// TIA Portal project "HydroPlantProject_V15.1" (V15.1)

(* hardware
DEVICE "S71500/ET200MP station_1"  S7-1500 station
   slot 0: "Rail_0"  Rack  6ES7 590-1***0-0AA0
   slot 1: "PLC_1"  CPU 1511-1 PN  6ES7 511-1AK00-0AB0  V1.8
      slot 3: "CPU display_1"  6ES7591-1AA00-0AA0
DEVICE "PC-System_1"  SIMATIC PC station
   slot 0: "SIMATIC PC station"  Rail  SIMATIC PC-Station  V1.0
      slot 125: "Stationmanager"  Station_Manager  V6.0.4
   slot 1: "HMI_RT_1"  WinCC RT Professional  6AV2 105-0xxxx-xxxx  15.1.0.0
   slot 2: "IE general_1"  IE General  IE_CP  V8.2.0
*)

// ===== PLC "PLC_1"  CPU 1511-1 PN =====

VAR_GLOBAL   // PLC tag table "Default tag table"
   "Brake_Out" AT %M4.0 : Bool;
   "OilPumpVFDsp_Out" AT %MW6 : Int;
   "OilTemp_In" AT %MW12 : Int;
   "kW_In" AT %MW14 : Int;
   "RPM_In" AT %MW16 : Int;
   "Baffle_Out" AT %MW18 : Int;
   "OilPumpVFDen_Out" AT %M4.1 : Bool;
   "ProgLang" AT %MW0 : Int;
   "ONS1" AT %M2.0 : Bool;
   "PB_LAD" AT %M2.1 : Bool;
   "ONS" AT %M2.2 : Bool;
   "ONS2" AT %M2.3 : Bool;
   "ONS3" AT %M2.4 : Bool;
   "PB_FBD" AT %M2.5 : Bool;
   "PB_SCL" AT %M2.6 : Bool;
   "PB_STL" AT %M2.7 : Bool;
   "AlarmHorn_Out" AT %M3.0 : Bool;
   "StationInterlock_Out" AT %M3.1 : Bool;
   "OilPumpVFDpct" AT %MW8 : Int;
   "BafflePct" AT %MW10 : Int;
   "OilTemp" AT %MW20 : Int;
   "OilFlow" AT %MW22 : Int;
   "OilFlow_In" AT %MW24 : Int;
   "RPM" AT %MW26 : Int;
   "Current" AT %MW28 : Int;
   "Current_In" AT %MW30 : Int;
   "OilPumpVFDoff_Pb" AT %M3.2 : Bool;
   "OilPumpVFDhand_Pb" AT %M3.3 : Bool;
   "OilPumpVFDauto_Pb" AT %M3.4 : Bool;
   "BrakeOff_Pb" AT %M3.5 : Bool;
   "BrakeHand_Pb" AT %M3.6 : Bool;
   "BrakeAuto_Pb" AT %M3.7 : Bool;
   "BrakeHoa" AT %MW34 : Int;
   "AlarmHornOff_Pb" AT %M4.2 : Bool;
   "AlarmHornHand_Pb" AT %M4.3 : Bool;
   "AlarmHornAuto_Pb" AT %M4.4 : Bool;
   "AlarmHornHoa" AT %MW36 : Int;
   "StationIntOff_Pb" AT %M4.5 : Bool;
   "StationIntHand_Pb" AT %M4.6 : Bool;
   "StationIntAuto_Pb" AT %M4.7 : Bool;
   "StationIntHoa" AT %MW38 : Int;
   "OilPumpVFD_Ctrl" AT %M5.0 : Bool;
   "StationIntl_Ctrl" AT %M5.1 : Bool;
   "AlarmHorn_Ctrl" AT %M5.2 : Bool;
   "Brake_Ctrl" AT %M5.3 : Bool;
   "OilLowFlowDelay_Sp" AT %MW40 : Int;
   "AlarmReset" AT %M5.4 : Bool;
   "AlarmSilence" AT %M5.5 : Bool;
   "OilLowFlowAlarm" AT %M5.6 : Bool;
   "OilLowFlowNotify" AT %M5.7 : Bool;
   "OilLLflowSp" AT %MW42 : Int;
   "OvercurrentDelay_Sp" AT %MW44 : Int;
   "OvercurrentSp" AT %MW46 : Int;
   "OvercurrentAlarm" AT %M48.0 : Bool;
   "OvercurrentNotify" AT %M48.1 : Bool;
   "HighOilTempDelay_Sp" AT %MW50 : Int;
   "HighOilTempAlarm" AT %M48.2 : Bool;
   "HighOilTempNotify" AT %M48.3 : Bool;
   "HighOilTempSp" AT %MW52 : Int;
   "OverspeedDelay_Sp" AT %MW54 : Int;
   "OverspeedSp" AT %MW56 : Int;
   "OverspeedAlarm" AT %M48.4 : Bool;
   "OverspeedNotify" AT %M48.5 : Bool;
   "OilHighFlowDelay_Sp" AT %MW58 : Int;
   "OilHHflowSp" AT %MW60 : Int;
   "OilHighFlowAlarm" AT %M48.6 : Bool;
   "OilHighFlowNotify" AT %M48.7 : Bool;
   "BrakeFailureDelay_Sp" AT %MW62 : Int;
   "BrakeFailureAlarm" AT %M49.0 : Bool;
   "BrakeFailureNotify" AT %M49.1 : Bool;
   "EStop" AT %M49.2 : Bool;
   "EStopAlarm" AT %M49.3 : Bool;
   "EStopNotify" AT %M49.4 : Bool;
   "Tag_1" AT %T1 : Timer;
   "Tag_2" AT %T2 : Timer;
   "ONS2(1)" AT %M49.5 : Bool;
   "ONS2(2)" AT %M49.6 : Bool;
   "Baffle_En" AT %M49.7 : Bool;
   "Deleteme" AT %M64.0 : Bool;
   "deleteme1" AT %MD66 : Real;
   "WarmupMode" AT %M64.1 : Bool;
   "StabilizeMode" AT %M64.2 : Bool;
   "GenerationMode" AT %M64.3 : Bool;
   "CooldownMode" AT %M64.4 : Bool;
   "IdleMode" AT %M64.5 : Bool;
   "FaultMode" AT %M64.6 : Bool;
   "WarmupRPM" AT %MW70 : Int;
   "BafflePIDSp" AT %MW72 : Int;
   "BaffleHOA" AT %MW74 : Int;
   "Baffle_Ctrl" AT %M64.7 : Bool;
   "VFD_Sp" AT %MW76 : Int;
   "WarmupVFDpct" AT %MW78 : Int;
   "WarmupOilTemp" AT %MW80 : Int;
   "WarmupOilTempDelaySp" AT %MW82 : Int;
   "WarmupTrasition" AT %M65.0 : Bool;
   "BafflePIDin" AT %MW84 : Int;
   "StabilizekWSp" AT %MW86 : Int;
   "StabilizeDelaySp" AT %MW88 : Int;
   "StabilizeTrasition" AT %M65.1 : Bool;
   "SystemStart_Pb" AT %M65.2 : Bool;
   "StartSequenceBit" AT %M65.3 : Bool;
   "SystemStop_Pb" AT %M65.4 : Bool;
   "GenerationTransition" AT %M65.5 : Bool;
   "CooldownRPM" AT %MW90 : Int;
   "CooldownDelaySp" AT %MW92 : Int;
   "CooldownTrasition" AT %M65.6 : Bool;
   "CooldownRPMSp" AT %MW94 : Int;
   "CooldownOilTempSp" AT %MW96 : Int;
   "ONS4" AT %M65.7 : Bool;
   "SequenceRunning" AT %M98.0 : Bool;
   "ONS5" AT %M98.1 : Bool;
   "HOFoverrideVFDsp" AT %MW100 : Int;
   "ONS6" AT %M98.2 : Bool;
   "BaffleManual" AT %M98.3 : Bool;
   "BaffleAuto_Pb" AT %M98.4 : Bool;
   "BaffleHand_Pb" AT %M98.5 : Bool;
   "BaffleOff_Pb" AT %M98.6 : Bool;
   "ONS8" AT %M98.7 : Bool;
   "BaffleManualSp" AT %MD102 : Real;
   "ONS9" AT %M99.0 : Bool;
   "ONS10" AT %M99.1 : Bool;
   "ONS7" AT %M99.2 : Bool;
   "VFDHand_Pb" AT %M99.3 : Bool;
   "VFDOff_Pb" AT %M99.4 : Bool;
   "VFDAuto_Pb" AT %M99.5 : Bool;
   "ONS11" AT %M99.6 : Bool;
   "ONS12" AT %M99.7 : Bool;
   "ONS13" AT %M106.0 : Bool;
   "VFDHOA" AT %MW108 : Int;
   "VFDManualSp" AT %MD110 : Real;
   "ONS14" AT %M106.1 : Bool;
   "ONS15" AT %M106.2 : Bool;
   "VFDmanual" AT %M106.3 : Bool;
   "OilPumpVFDon" AT %M106.4 : Bool;
   "BafflePID_On" AT %M106.5 : Bool;
   "FullAutoBit" AT %M106.6 : Bool;
   "HM_Minutes" AT %MW32 : Int;
   "HM_Hours" AT %MW114 : Int;
   "HM_Days" AT %MW116 : Int;
   "ResetHourmeter_Pb" AT %M106.7 : Bool;
   "ModeInt" AT %MW118 : Int;
END_VAR

DATA_BLOCK "SimLogic_DB"   // DB1
{ S7_Optimized_Access := 'TRUE' }
VERSION : 0.1
// stored: InstanceOfName SimLogic
"SimLogic"
BEGIN
END_DATA_BLOCK

DATA_BLOCK "MODES_LAD_DB"   // DB2
{ S7_Optimized_Access := 'TRUE' }
VERSION : 0.1
// stored: InstanceOfName MODES_LAD
"MODES_LAD"
BEGIN
END_DATA_BLOCK

DATA_BLOCK "MODES_FBD_DB"   // DB4
{ S7_Optimized_Access := 'TRUE' }
VERSION : 0.1
// stored: InstanceOfName MODES_FBD
"MODES_FBD"
BEGIN
END_DATA_BLOCK

DATA_BLOCK "IO_LAD_DB"   // DB5
{ S7_Optimized_Access := 'TRUE' }
VERSION : 0.1
// stored: InstanceOfName IO_LAD
"IO_LAD"
BEGIN
END_DATA_BLOCK

DATA_BLOCK "IO_FBD_DB"   // DB6
{ S7_Optimized_Access := 'TRUE' }
VERSION : 0.1
// stored: InstanceOfName IO_FBD
"IO_FBD"
BEGIN
END_DATA_BLOCK

DATA_BLOCK "IO_SCL_DB"   // DB7
{ S7_Optimized_Access := 'TRUE' }
VERSION : 0.1
// stored: InstanceOfName IO_SCL
"IO_SCL"
BEGIN
END_DATA_BLOCK

DATA_BLOCK "IO_STL_DB"   // DB8
{ S7_Optimized_Access := 'TRUE' }
VERSION : 0.1
// stored: InstanceOfName IO_STL
"IO_STL"
BEGIN
END_DATA_BLOCK

DATA_BLOCK "ALARMS_LAD_DB"   // DB9
{ S7_Optimized_Access := 'TRUE' }
VERSION : 0.1
// stored: InstanceOfName ALARMS_LAD
"ALARMS_LAD"
BEGIN
END_DATA_BLOCK

DATA_BLOCK "HOA_LAD_DB"   // DB10
{ S7_Optimized_Access := 'TRUE' }
VERSION : 0.1
// stored: InstanceOfName HOA_LAD
"HOA_LAD"
BEGIN
END_DATA_BLOCK

DATA_BLOCK "HOA_FBD_DB"   // DB11
{ S7_Optimized_Access := 'TRUE' }
VERSION : 0.1
// stored: InstanceOfName HOA_FBD
"HOA_FBD"
BEGIN
END_DATA_BLOCK

DATA_BLOCK "HOA_SCL_DB"   // DB12
{ S7_Optimized_Access := 'TRUE' }
VERSION : 0.1
// stored: InstanceOfName HOA_SCL
"HOA_SCL"
BEGIN
END_DATA_BLOCK

DATA_BLOCK "HOA_STL_DB"   // DB13
{ S7_Optimized_Access := 'TRUE' }
VERSION : 0.1
// stored: InstanceOfName HOA_STL
"HOA_STL"
BEGIN
END_DATA_BLOCK

DATA_BLOCK "ALARMS_FBD_DB"   // DB14
{ S7_Optimized_Access := 'TRUE' }
VERSION : 0.1
// stored: InstanceOfName ALARMS_FBD
"ALARMS_FBD"
BEGIN
END_DATA_BLOCK

DATA_BLOCK "ALARMS_SCL_DB"   // DB15
{ S7_Optimized_Access := 'TRUE' }
VERSION : 0.1
// stored: InstanceOfName ALARMS_SCL
"ALARMS_SCL"
BEGIN
END_DATA_BLOCK

DATA_BLOCK "ALARMS_STL_DB"   // DB16
{ S7_Optimized_Access := 'TRUE' }
VERSION : 0.1
// stored: InstanceOfName ALARMS_STL
"ALARMS_STL"
BEGIN
END_DATA_BLOCK

DATA_BLOCK "MODES_SCL_DB"   // DB44
{ S7_Optimized_Access := 'TRUE' }
VERSION : 0.1
// stored: InstanceOfName MODES_SCL
"MODES_SCL"
BEGIN
END_DATA_BLOCK

DATA_BLOCK "MODES_STL_DB"   // DB45
{ S7_Optimized_Access := 'TRUE' }
VERSION : 0.1
// stored: InstanceOfName MODES_STL
"MODES_STL"
BEGIN
END_DATA_BLOCK

DATA_BLOCK "SEQUENCE_DB"   // DB58
{ S7_Optimized_Access := 'TRUE' }
VERSION : 0.1
// stored: InstanceOfName SEQUENCE
"SEQUENCE"
BEGIN
END_DATA_BLOCK

DATA_BLOCK "HOURMETER_LAD_DB"   // DB61
{ S7_Optimized_Access := 'TRUE' }
VERSION : 0.1
// stored: InstanceOfName HOURMETER_LAD
"HOURMETER_LAD"
BEGIN
END_DATA_BLOCK

DATA_BLOCK "HOURMETER_FBD_DB"   // DB62
{ S7_Optimized_Access := 'TRUE' }
VERSION : 0.1
// stored: InstanceOfName HOURMETER_FBD
"HOURMETER_FBD"
BEGIN
END_DATA_BLOCK

DATA_BLOCK "HOURMETER_SCL_DB"   // DB63
{ S7_Optimized_Access := 'TRUE' }
VERSION : 0.1
// stored: InstanceOfName HOURMETER_SCL
"HOURMETER_SCL"
BEGIN
END_DATA_BLOCK

DATA_BLOCK "HOURMETER_STL_DB"   // DB64
{ S7_Optimized_Access := 'TRUE' }
VERSION : 0.1
// stored: InstanceOfName HOURMETER_STL
"HOURMETER_STL"
BEGIN
END_DATA_BLOCK

// folder: System blocks/Program resources

DATA_BLOCK "IEC_Timer_0_DB_25"   // DB3
{ S7_Optimized_Access := 'TRUE' }
AUTHOR : Simatic
FAMILY : IEC
NAME : IEC_TMR
VERSION : 1.0
// stored: InstanceOfName IEC_TIMER
"IEC_TIMER"
BEGIN
END_DATA_BLOCK

DATA_BLOCK "IEC_Timer_0_DB"   // DB17
{ S7_Optimized_Access := 'TRUE' }
AUTHOR : Simatic
FAMILY : IEC
NAME : IEC_TMR
VERSION : 1.0
// stored: InstanceOfName IEC_TIMER
"IEC_TIMER"
BEGIN
END_DATA_BLOCK

DATA_BLOCK "IEC_Timer_0_DB_1"   // DB18
{ S7_Optimized_Access := 'TRUE' }
AUTHOR : Simatic
FAMILY : IEC
NAME : IEC_TMR
VERSION : 1.0
// stored: InstanceOfName IEC_TIMER
"IEC_TIMER"
BEGIN
END_DATA_BLOCK

DATA_BLOCK "IEC_Timer_0_DB_2"   // DB19
{ S7_Optimized_Access := 'TRUE' }
AUTHOR : Simatic
FAMILY : IEC
NAME : IEC_TMR
VERSION : 1.0
// stored: InstanceOfName IEC_TIMER
"IEC_TIMER"
BEGIN
END_DATA_BLOCK

DATA_BLOCK "IEC_Timer_0_DB_3"   // DB20
{ S7_Optimized_Access := 'TRUE' }
AUTHOR : Simatic
FAMILY : IEC
NAME : IEC_TMR
VERSION : 1.0
// stored: InstanceOfName IEC_TIMER
"IEC_TIMER"
BEGIN
END_DATA_BLOCK

DATA_BLOCK "IEC_Timer_0_DB_4"   // DB21
{ S7_Optimized_Access := 'TRUE' }
AUTHOR : Simatic
FAMILY : IEC
NAME : IEC_TMR
VERSION : 1.0
// stored: InstanceOfName IEC_TIMER
"IEC_TIMER"
BEGIN
END_DATA_BLOCK

DATA_BLOCK "IEC_Timer_0_DB_5"   // DB22
{ S7_Optimized_Access := 'TRUE' }
AUTHOR : Simatic
FAMILY : IEC
NAME : IEC_TMR
VERSION : 1.0
// stored: InstanceOfName IEC_TIMER
"IEC_TIMER"
BEGIN
END_DATA_BLOCK

DATA_BLOCK "IEC_Timer_0_DB_6"   // DB23
{ S7_Optimized_Access := 'TRUE' }
AUTHOR : Simatic
FAMILY : IEC
NAME : IEC_TMR
VERSION : 1.0
// stored: InstanceOfName IEC_TIMER
"IEC_TIMER"
BEGIN
END_DATA_BLOCK

DATA_BLOCK "IEC_Timer_0_DB_7"   // DB24
{ S7_Optimized_Access := 'TRUE' }
AUTHOR : Simatic
FAMILY : IEC
NAME : IEC_TMR
VERSION : 1.0
// stored: InstanceOfName IEC_TIMER
"IEC_TIMER"
BEGIN
END_DATA_BLOCK

DATA_BLOCK "IEC_Timer_0_DB_8"   // DB25
{ S7_Optimized_Access := 'TRUE' }
AUTHOR : Simatic
FAMILY : IEC
NAME : IEC_TMR
VERSION : 1.0
// stored: InstanceOfName IEC_TIMER
"IEC_TIMER"
BEGIN
END_DATA_BLOCK

DATA_BLOCK "IEC_Timer_0_DB_9"   // DB26
{ S7_Optimized_Access := 'TRUE' }
AUTHOR : Simatic
FAMILY : IEC
NAME : IEC_TMR
VERSION : 1.0
// stored: InstanceOfName IEC_TIMER
"IEC_TIMER"
BEGIN
END_DATA_BLOCK

DATA_BLOCK "IEC_Timer_0_DB_10"   // DB27
{ S7_Optimized_Access := 'TRUE' }
AUTHOR : Simatic
FAMILY : IEC
NAME : IEC_TMR
VERSION : 1.0
// stored: InstanceOfName IEC_TIMER
"IEC_TIMER"
BEGIN
END_DATA_BLOCK

DATA_BLOCK "IEC_Timer_0_DB_110"   // DB28
{ S7_Optimized_Access := 'TRUE' }
AUTHOR : Simatic
FAMILY : IEC
NAME : IEC_TMR
VERSION : 1.0
// stored: InstanceOfName IEC_TIMER
"IEC_TIMER"
BEGIN
END_DATA_BLOCK

DATA_BLOCK "IEC_Timer_0_DB_11"   // DB29
{ S7_Optimized_Access := 'TRUE' }
AUTHOR : Simatic
FAMILY : IEC
NAME : IEC_TMR
VERSION : 1.0
// stored: InstanceOfName IEC_TIMER
"IEC_TIMER"
BEGIN
END_DATA_BLOCK

DATA_BLOCK "IEC_Timer_0_DB_12"   // DB30
{ S7_Optimized_Access := 'TRUE' }
AUTHOR : Simatic
FAMILY : IEC
NAME : IEC_TMR
VERSION : 1.0
// stored: InstanceOfName IEC_TIMER
"IEC_TIMER"
BEGIN
END_DATA_BLOCK

DATA_BLOCK "IEC_Timer_0_DB_13"   // DB31
{ S7_Optimized_Access := 'TRUE' }
AUTHOR : Simatic
FAMILY : IEC
NAME : IEC_TMR
VERSION : 1.0
// stored: InstanceOfName IEC_TIMER
"IEC_TIMER"
BEGIN
END_DATA_BLOCK

DATA_BLOCK "IEC_Timer_0_DB_14"   // DB32
{ S7_Optimized_Access := 'TRUE' }
AUTHOR : Simatic
FAMILY : IEC
NAME : IEC_TMR
VERSION : 1.0
// stored: InstanceOfName IEC_TIMER
"IEC_TIMER"
BEGIN
END_DATA_BLOCK

DATA_BLOCK "IEC_Timer_0_DB_15"   // DB33
{ S7_Optimized_Access := 'TRUE' }
AUTHOR : Simatic
FAMILY : IEC
NAME : IEC_TMR
VERSION : 1.0
// stored: InstanceOfName IEC_TIMER
"IEC_TIMER"
BEGIN
END_DATA_BLOCK

DATA_BLOCK "IEC_Timer_0_DB_16"   // DB34
{ S7_Optimized_Access := 'TRUE' }
AUTHOR : Simatic
FAMILY : IEC
NAME : IEC_TMR
VERSION : 1.0
// stored: InstanceOfName IEC_TIMER
"IEC_TIMER"
BEGIN
END_DATA_BLOCK

DATA_BLOCK "IEC_Timer_0_DB_17"   // DB35
{ S7_Optimized_Access := 'TRUE' }
AUTHOR : Simatic
FAMILY : IEC
NAME : IEC_TMR
VERSION : 1.0
// stored: InstanceOfName IEC_TIMER
"IEC_TIMER"
BEGIN
END_DATA_BLOCK

DATA_BLOCK "IEC_Timer_0_DB_18"   // DB36
{ S7_Optimized_Access := 'TRUE' }
AUTHOR : Simatic
FAMILY : IEC
NAME : IEC_TMR
VERSION : 1.0
// stored: InstanceOfName IEC_TIMER
"IEC_TIMER"
BEGIN
END_DATA_BLOCK

DATA_BLOCK "IEC_Timer_0_DB_19"   // DB37
{ S7_Optimized_Access := 'TRUE' }
AUTHOR : Simatic
FAMILY : IEC
NAME : IEC_TMR
VERSION : 1.0
// stored: InstanceOfName IEC_TIMER
"IEC_TIMER"
BEGIN
END_DATA_BLOCK

DATA_BLOCK "IEC_Timer_0_DB_20"   // DB38
{ S7_Optimized_Access := 'TRUE' }
AUTHOR : Simatic
FAMILY : IEC
NAME : IEC_TMR
VERSION : 1.0
// stored: InstanceOfName IEC_TIMER
"IEC_TIMER"
BEGIN
END_DATA_BLOCK

DATA_BLOCK "IEC_Timer_0_DB_21"   // DB39
{ S7_Optimized_Access := 'TRUE' }
AUTHOR : Simatic
FAMILY : IEC
NAME : IEC_TMR
VERSION : 1.0
// stored: InstanceOfName IEC_TIMER
"IEC_TIMER"
BEGIN
END_DATA_BLOCK

DATA_BLOCK "IEC_Timer_0_DB_22"   // DB40
{ S7_Optimized_Access := 'TRUE' }
AUTHOR : Simatic
FAMILY : IEC
NAME : IEC_TMR
VERSION : 1.0
// stored: InstanceOfName IEC_TIMER
"IEC_TIMER"
BEGIN
END_DATA_BLOCK

DATA_BLOCK "IEC_Timer_0_DB_23"   // DB41
{ S7_Optimized_Access := 'TRUE' }
AUTHOR : Simatic
FAMILY : IEC
NAME : IEC_TMR
VERSION : 1.0
// stored: InstanceOfName IEC_TIMER
"IEC_TIMER"
BEGIN
END_DATA_BLOCK

DATA_BLOCK "IEC_Timer_1_DB"   // DB43
{ S7_Optimized_Access := 'TRUE' }
AUTHOR : Simatic
FAMILY : IEC
NAME : IEC_TMR
VERSION : 1.0
// stored: InstanceOfName IEC_TIMER
"IEC_TIMER"
BEGIN
END_DATA_BLOCK

DATA_BLOCK "IEC_Timer_0_DB_24"   // DB46
{ S7_Optimized_Access := 'TRUE' }
AUTHOR : Simatic
FAMILY : IEC
NAME : IEC_TMR
VERSION : 1.0
// stored: InstanceOfName IEC_TIMER
"IEC_TIMER"
BEGIN
END_DATA_BLOCK

DATA_BLOCK "IEC_Timer_0_DB_26"   // DB47
{ S7_Optimized_Access := 'TRUE' }
AUTHOR : Simatic
FAMILY : IEC
NAME : IEC_TMR
VERSION : 1.0
// stored: InstanceOfName IEC_TIMER
"IEC_TIMER"
BEGIN
END_DATA_BLOCK

DATA_BLOCK "IEC_Timer_0_DB_27"   // DB48
{ S7_Optimized_Access := 'TRUE' }
AUTHOR : Simatic
FAMILY : IEC
NAME : IEC_TMR
VERSION : 1.0
// stored: InstanceOfName IEC_TIMER
"IEC_TIMER"
BEGIN
END_DATA_BLOCK

DATA_BLOCK "IEC_Timer_0_DB_28"   // DB49
{ S7_Optimized_Access := 'TRUE' }
AUTHOR : Simatic
FAMILY : IEC
NAME : IEC_TMR
VERSION : 1.0
// stored: InstanceOfName IEC_TIMER
"IEC_TIMER"
BEGIN
END_DATA_BLOCK

DATA_BLOCK "IEC_Timer_0_DB_29"   // DB50
{ S7_Optimized_Access := 'TRUE' }
AUTHOR : Simatic
FAMILY : IEC
NAME : IEC_TMR
VERSION : 1.0
// stored: InstanceOfName IEC_TIMER
"IEC_TIMER"
BEGIN
END_DATA_BLOCK

DATA_BLOCK "IEC_Timer_0_DB_30"   // DB51
{ S7_Optimized_Access := 'TRUE' }
AUTHOR : Simatic
FAMILY : IEC
NAME : IEC_TMR
VERSION : 1.0
// stored: InstanceOfName IEC_TIMER
"IEC_TIMER"
BEGIN
END_DATA_BLOCK

DATA_BLOCK "IEC_Timer_0_DB_31"   // DB52
{ S7_Optimized_Access := 'TRUE' }
AUTHOR : Simatic
FAMILY : IEC
NAME : IEC_TMR
VERSION : 1.0
// stored: InstanceOfName IEC_TIMER
"IEC_TIMER"
BEGIN
END_DATA_BLOCK

DATA_BLOCK "IEC_Timer_0_DB_32"   // DB53
{ S7_Optimized_Access := 'TRUE' }
AUTHOR : Simatic
FAMILY : IEC
NAME : IEC_TMR
VERSION : 1.0
// stored: InstanceOfName IEC_TIMER
"IEC_TIMER"
BEGIN
END_DATA_BLOCK

DATA_BLOCK "IEC_Timer_0_DB_33"   // DB54
{ S7_Optimized_Access := 'TRUE' }
AUTHOR : Simatic
FAMILY : IEC
NAME : IEC_TMR
VERSION : 1.0
// stored: InstanceOfName IEC_TIMER
"IEC_TIMER"
BEGIN
END_DATA_BLOCK

DATA_BLOCK "IEC_Timer_0_DB_34"   // DB55
{ S7_Optimized_Access := 'TRUE' }
AUTHOR : Simatic
FAMILY : IEC
NAME : IEC_TMR
VERSION : 1.0
// stored: InstanceOfName IEC_TIMER
"IEC_TIMER"
BEGIN
END_DATA_BLOCK

DATA_BLOCK "IEC_Timer_0_DB_35"   // DB56
{ S7_Optimized_Access := 'TRUE' }
AUTHOR : Simatic
FAMILY : IEC
NAME : IEC_TMR
VERSION : 1.0
// stored: InstanceOfName IEC_TIMER
"IEC_TIMER"
BEGIN
END_DATA_BLOCK

DATA_BLOCK "IEC_Timer_0_DB_36"   // DB57
{ S7_Optimized_Access := 'TRUE' }
AUTHOR : Simatic
FAMILY : IEC
NAME : IEC_TMR
VERSION : 1.0
// stored: InstanceOfName IEC_TIMER
"IEC_TIMER"
BEGIN
END_DATA_BLOCK

DATA_BLOCK "IEC_Timer_0_DB_37"   // DB65
{ S7_Optimized_Access := 'TRUE' }
AUTHOR : Simatic
FAMILY : IEC
NAME : IEC_TMR
VERSION : 1.0
// stored: InstanceOfName IEC_TIMER
"IEC_TIMER"
BEGIN
END_DATA_BLOCK

DATA_BLOCK "IEC_Counter_0_DB"   // DB66
{ S7_Optimized_Access := 'TRUE' }
AUTHOR : Simatic
FAMILY : IEC
NAME : CNTR
VERSION : 1.0
// stored: InstanceOfName IEC_COUNTER
"IEC_COUNTER"
BEGIN
END_DATA_BLOCK

DATA_BLOCK "IEC_Counter_0_DB_1"   // DB67
{ S7_Optimized_Access := 'TRUE' }
AUTHOR : Simatic
FAMILY : IEC
NAME : CNTR
VERSION : 1.0
// stored: InstanceOfName IEC_COUNTER
"IEC_COUNTER"
BEGIN
END_DATA_BLOCK

DATA_BLOCK "IEC_Counter_0_DB_2"   // DB68
{ S7_Optimized_Access := 'TRUE' }
AUTHOR : Simatic
FAMILY : IEC
NAME : CNTR
VERSION : 1.0
// stored: InstanceOfName IEC_COUNTER
"IEC_COUNTER"
BEGIN
END_DATA_BLOCK

DATA_BLOCK "IEC_Timer_0_DB_38"   // DB69
{ S7_Optimized_Access := 'TRUE' }
AUTHOR : Simatic
FAMILY : IEC
NAME : IEC_TMR
VERSION : 1.0
// stored: InstanceOfName IEC_TIMER
"IEC_TIMER"
BEGIN
END_DATA_BLOCK

DATA_BLOCK "IEC_Timer_0_DB_39"   // DB70
{ S7_Optimized_Access := 'TRUE' }
AUTHOR : Simatic
FAMILY : IEC
NAME : IEC_TMR
VERSION : 1.0
// stored: InstanceOfName IEC_TIMER
"IEC_TIMER"
BEGIN
END_DATA_BLOCK

DATA_BLOCK "IEC_Timer_0_DB_40"   // DB71
{ S7_Optimized_Access := 'TRUE' }
AUTHOR : Simatic
FAMILY : IEC
NAME : IEC_TMR
VERSION : 1.0
// stored: InstanceOfName IEC_TIMER
"IEC_TIMER"
BEGIN
END_DATA_BLOCK

DATA_BLOCK "IEC_Counter_0_DB_3"   // DB72
{ S7_Optimized_Access := 'TRUE' }
AUTHOR : Simatic
FAMILY : IEC
NAME : CNTR
VERSION : 1.0
// stored: InstanceOfName IEC_COUNTER
"IEC_COUNTER"
BEGIN
END_DATA_BLOCK

DATA_BLOCK "IEC_Counter_0_DB_4"   // DB73
{ S7_Optimized_Access := 'TRUE' }
AUTHOR : Simatic
FAMILY : IEC
NAME : CNTR
VERSION : 1.0
// stored: InstanceOfName IEC_COUNTER
"IEC_COUNTER"
BEGIN
END_DATA_BLOCK

DATA_BLOCK "IEC_Counter_0_DB_5"   // DB74
{ S7_Optimized_Access := 'TRUE' }
AUTHOR : Simatic
FAMILY : IEC
NAME : CNTR
VERSION : 1.0
// stored: InstanceOfName IEC_COUNTER
"IEC_COUNTER"
BEGIN
END_DATA_BLOCK

DATA_BLOCK "IEC_Timer_0_DB_41"   // DB75
{ S7_Optimized_Access := 'TRUE' }
AUTHOR : Simatic
FAMILY : IEC
NAME : IEC_TMR
VERSION : 1.0
// stored: InstanceOfName IEC_TIMER
"IEC_TIMER"
BEGIN
END_DATA_BLOCK

DATA_BLOCK "IEC_Counter_0_DB_6"   // DB76
{ S7_Optimized_Access := 'TRUE' }
AUTHOR : Simatic
FAMILY : IEC
NAME : CNTR
VERSION : 1.0
// stored: InstanceOfName IEC_COUNTER
"IEC_COUNTER"
BEGIN
END_DATA_BLOCK

DATA_BLOCK "IEC_Counter_0_DB_7"   // DB77
{ S7_Optimized_Access := 'TRUE' }
AUTHOR : Simatic
FAMILY : IEC
NAME : CNTR
VERSION : 1.0
// stored: InstanceOfName IEC_COUNTER
"IEC_COUNTER"
BEGIN
END_DATA_BLOCK

DATA_BLOCK "IEC_Counter_0_DB_9"   // DB79
{ S7_Optimized_Access := 'TRUE' }
AUTHOR : Simatic
FAMILY : IEC
NAME : CNTR
VERSION : 1.0
// stored: InstanceOfName IEC_COUNTER
"IEC_COUNTER"
BEGIN
END_DATA_BLOCK

DATA_BLOCK "IEC_Timer_0_DB_42"   // DB80
{ S7_Optimized_Access := 'TRUE' }
AUTHOR : Simatic
FAMILY : IEC
NAME : IEC_TMR
VERSION : 1.0
// stored: InstanceOfName IEC_TIMER
"IEC_TIMER"
BEGIN
END_DATA_BLOCK

DATA_BLOCK "IEC_Timer_0_DB_43"   // DB81
{ S7_Optimized_Access := 'TRUE' }
AUTHOR : Simatic
FAMILY : IEC
NAME : IEC_TMR
VERSION : 1.0
// stored: InstanceOfName IEC_TIMER
"IEC_TIMER"
BEGIN
END_DATA_BLOCK

DATA_BLOCK "IEC_Counter_0_DB_10"   // DB82
{ S7_Optimized_Access := 'TRUE' }
AUTHOR : Simatic
FAMILY : IEC
NAME : CNTR
VERSION : 1.0
// stored: InstanceOfName IEC_COUNTER
"IEC_COUNTER"
BEGIN
END_DATA_BLOCK

DATA_BLOCK "IEC_Counter_0_DB_11"   // DB83
{ S7_Optimized_Access := 'TRUE' }
AUTHOR : Simatic
FAMILY : IEC
NAME : CNTR
VERSION : 1.0
// stored: InstanceOfName IEC_COUNTER
"IEC_COUNTER"
BEGIN
END_DATA_BLOCK

DATA_BLOCK "IEC_Counter_0_DB_12"   // DB84
{ S7_Optimized_Access := 'TRUE' }
AUTHOR : Simatic
FAMILY : IEC
NAME : CNTR
VERSION : 1.0
// stored: InstanceOfName IEC_COUNTER
"IEC_COUNTER"
BEGIN
END_DATA_BLOCK

DATA_BLOCK "IEC_Timer_0_DB_44"   // DB85
{ S7_Optimized_Access := 'TRUE' }
AUTHOR : Simatic
FAMILY : IEC
NAME : IEC_TMR
VERSION : 1.0
// stored: InstanceOfName IEC_TIMER
"IEC_TIMER"
BEGIN
END_DATA_BLOCK

// folder: (top level)

FUNCTION_BLOCK "SimLogic"   // FB1, FBD
{ S7_Optimized_Access := 'TRUE' }
VERSION : 0.1
   VAR
      "TO" : Bool;
      rpmv : Int;
      addrpmv : Bool;
      otsp : Int;
      ott : Int;
      TO1 : Bool;
      TO2 : Bool;
      be2 : Int;
      be3 : Int;
      be1 : Int;
      TO3 : Bool;
   END_VAR
   VAR_TEMP
      bf : Int;
      rpmvt : Int;
      bfr : Real;
   END_VAR
BEGIN

REGION Network 1
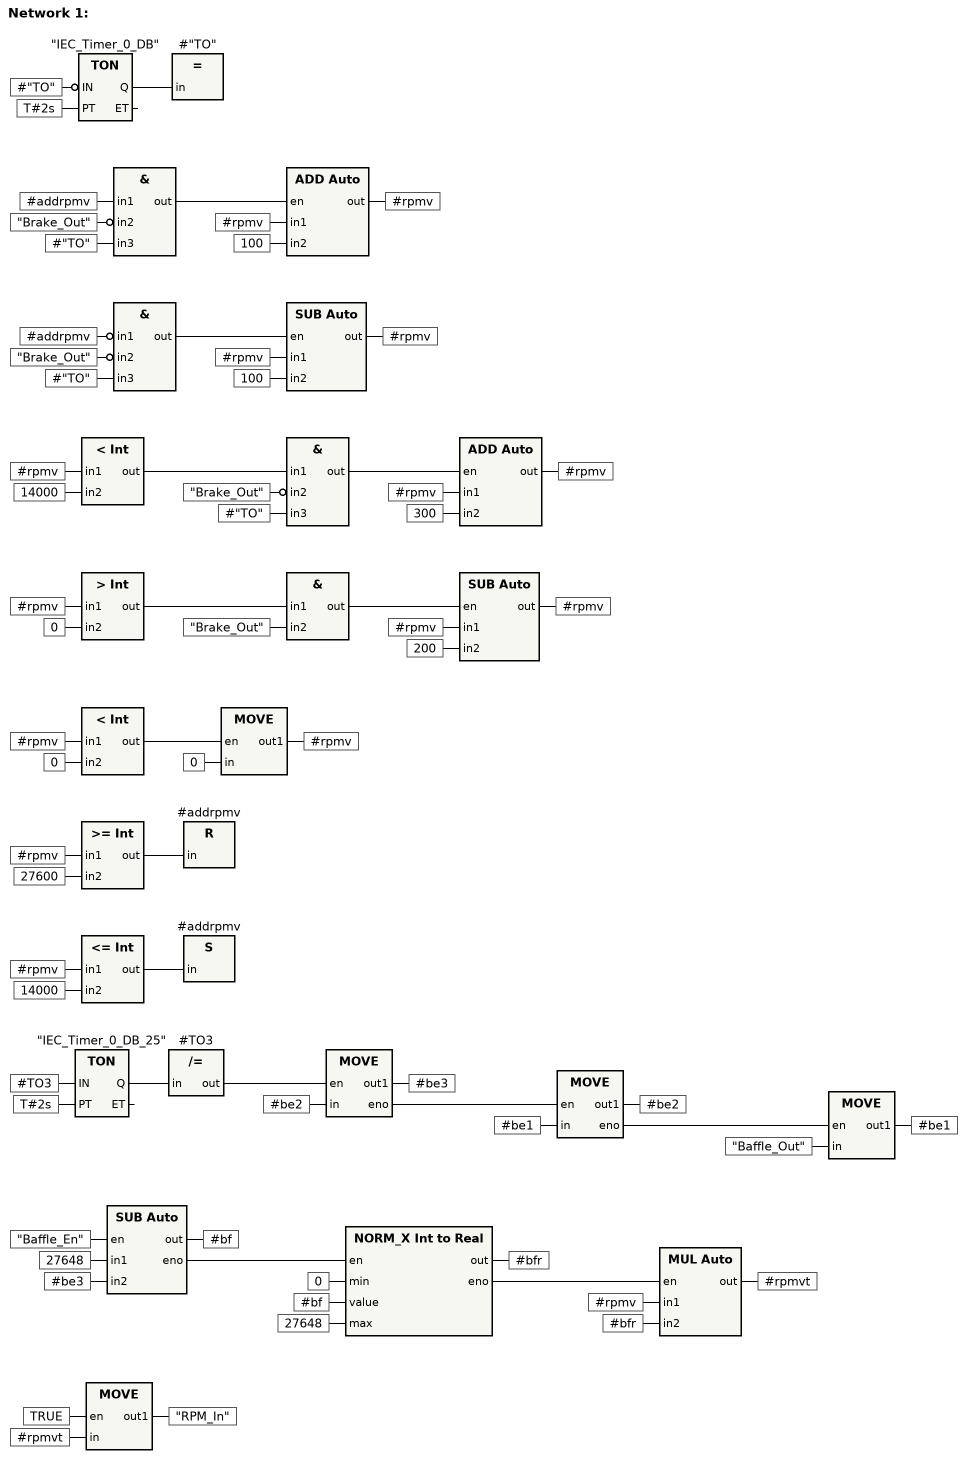
   "IEC_Timer_0_DB".TON(IN := NOT #"TO", PT := T#2s);
   #"TO" := "IEC_Timer_0_DB".Q;
   IF #addrpmv AND NOT "Brake_Out" AND #"TO" THEN #rpmv := #rpmv + 100; END_IF;
   IF NOT #addrpmv AND NOT "Brake_Out" AND #"TO" THEN #rpmv := #rpmv - 100; END_IF;
   IF (#rpmv < 14000) AND NOT "Brake_Out" AND #"TO" THEN #rpmv := #rpmv + 300; END_IF;
   IF (#rpmv > 0) AND "Brake_Out" THEN #rpmv := #rpmv - 200; END_IF;
   IF #rpmv < 0 THEN #rpmv := 0; END_IF;
   IF #rpmv >= 27600 THEN #addrpmv := FALSE; END_IF;
   IF #rpmv <= 14000 THEN #addrpmv := TRUE; END_IF;
   "IEC_Timer_0_DB_25".TON(IN := #TO3, PT := T#2s);
   #TO3 := NOT "IEC_Timer_0_DB_25".Q;
   IF "IEC_Timer_0_DB_25".Q THEN
       #be3 := #be2;
       #be2 := #be1;
       #be1 := "Baffle_Out";
   END_IF;
   IF "Baffle_En" THEN
       #bf := 27648 - #be3;
       #bfr := NORM_X(MIN := 0, VALUE := #bf, MAX := 27648);
       #rpmvt := #rpmv * #bfr;
   END_IF;
   IF TRUE THEN "RPM_In" := #rpmvt; END_IF;
END_REGION

REGION Network 2
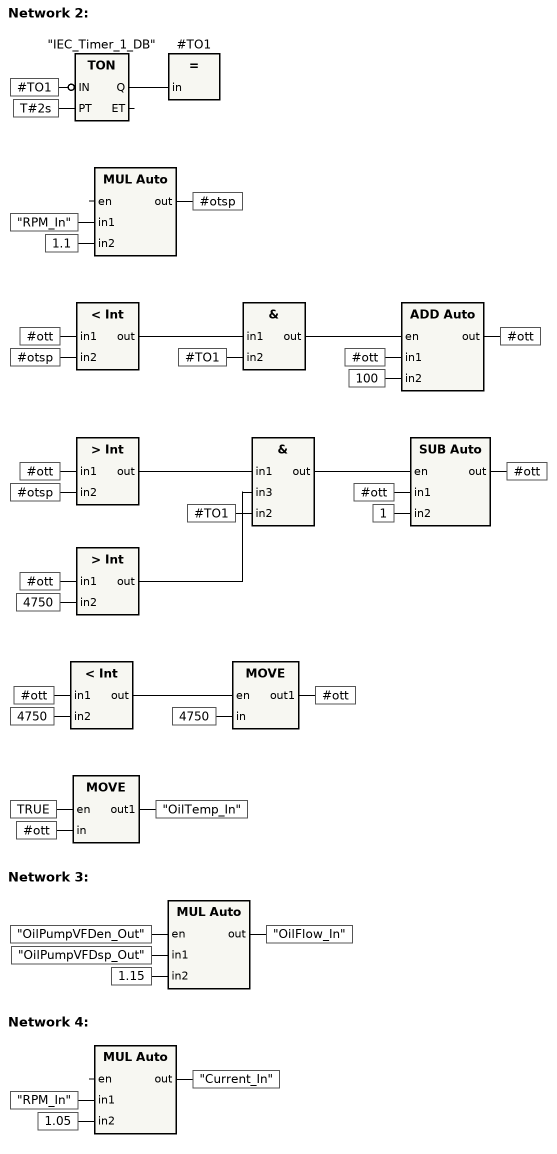
   "IEC_Timer_1_DB".TON(IN := NOT #TO1, PT := T#2s);
   #TO1 := "IEC_Timer_1_DB".Q;
   #otsp := "RPM_In" * 1.1;
   IF (#ott < #otsp) AND #TO1 THEN #ott := #ott + 100; END_IF;
   IF (#ott > #otsp) AND (#ott > 4750) AND #TO1 THEN #ott := #ott - 1; END_IF;
   IF #ott < 4750 THEN #ott := 4750; END_IF;
   IF TRUE THEN "OilTemp_In" := #ott; END_IF;
END_REGION

REGION Network 3
   IF "OilPumpVFDen_Out" THEN "OilFlow_In" := "OilPumpVFDsp_Out" * 1.15; END_IF;
END_REGION

REGION Network 4
   "Current_In" := "RPM_In" * 1.05;
END_REGION
END_FUNCTION_BLOCK

FUNCTION_BLOCK "IO_LAD"   // FB2, LAD
{ S7_Optimized_Access := 'TRUE' }
VERSION : 0.1
BEGIN

REGION Network 1
   // Digital Output
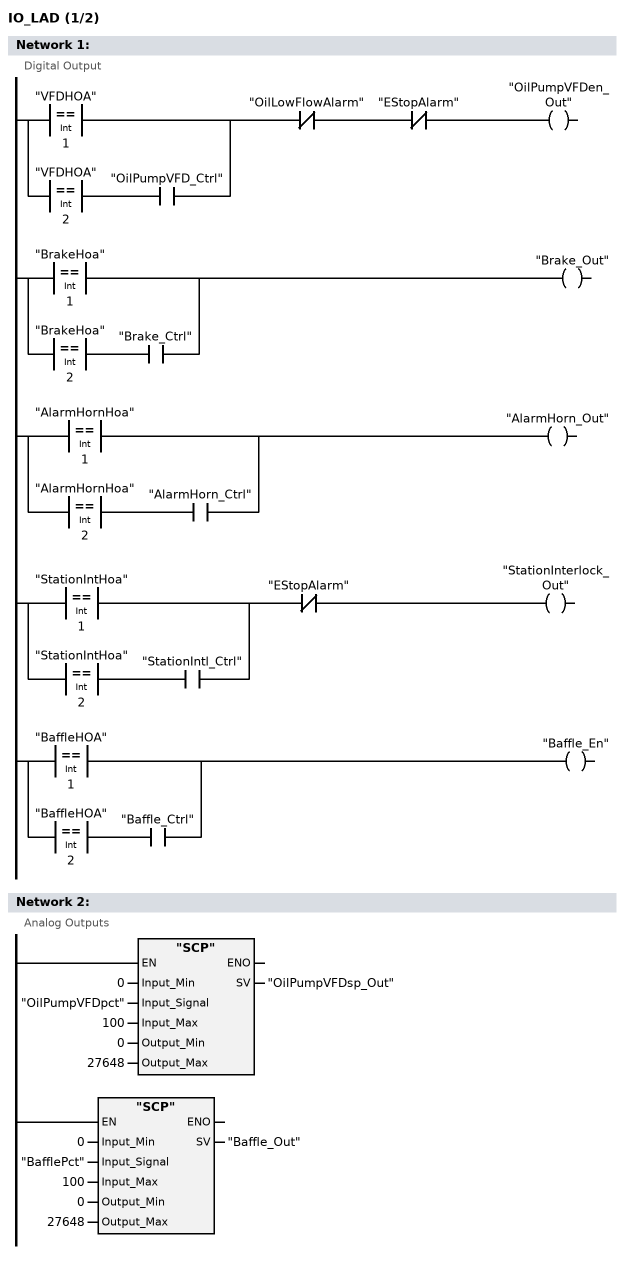
   RUNG wire#powerrail
      { S7_Templates := "SrcType := Int" } EQ_Contact(in1 := "VFDHOA", in2 := 1)
      wire#w1
      I_Contact( "OilLowFlowAlarm" )
      I_Contact( "EStopAlarm" )
      Coil( "OilPumpVFDen_Out" )
   END_RUNG
   RUNG wire#powerrail
      { S7_Templates := "SrcType := Int" } EQ_Contact(in1 := "VFDHOA", in2 := 2)
      Contact( "OilPumpVFD_Ctrl" )
   END_RUNG wire#w1
   RUNG wire#powerrail
      { S7_Templates := "SrcType := Int" } EQ_Contact(in1 := "BrakeHoa", in2 := 1)
      wire#w2
      Coil( "Brake_Out" )
   END_RUNG
   RUNG wire#powerrail
      { S7_Templates := "SrcType := Int" } EQ_Contact(in1 := "BrakeHoa", in2 := 2)
      Contact( "Brake_Ctrl" )
   END_RUNG wire#w2
   RUNG wire#powerrail
      { S7_Templates := "SrcType := Int" } EQ_Contact(in1 := "AlarmHornHoa", in2 := 1)
      wire#w3
      Coil( "AlarmHorn_Out" )
   END_RUNG
   RUNG wire#powerrail
      { S7_Templates := "SrcType := Int" } EQ_Contact(in1 := "AlarmHornHoa", in2 := 2)
      Contact( "AlarmHorn_Ctrl" )
   END_RUNG wire#w3
   RUNG wire#powerrail
      { S7_Templates := "SrcType := Int" } EQ_Contact(in1 := "StationIntHoa", in2 := 1)
      wire#w4
      I_Contact( "EStopAlarm" )
      Coil( "StationInterlock_Out" )
   END_RUNG
   RUNG wire#powerrail
      { S7_Templates := "SrcType := Int" } EQ_Contact(in1 := "StationIntHoa", in2 := 2)
      Contact( "StationIntl_Ctrl" )
   END_RUNG wire#w4
   RUNG wire#powerrail
      { S7_Templates := "SrcType := Int" } EQ_Contact(in1 := "BaffleHOA", in2 := 1)
      wire#w5
      Coil( "Baffle_En" )
   END_RUNG
   RUNG wire#powerrail
      { S7_Templates := "SrcType := Int" } EQ_Contact(in1 := "BaffleHOA", in2 := 2)
      Contact( "Baffle_Ctrl" )
   END_RUNG wire#w5
   // the same network as SCL:
   "OilPumpVFDen_Out" := (("VFDHOA" = 1) OR (("VFDHOA" = 2) AND "OilPumpVFD_Ctrl")) AND NOT "OilLowFlowAlarm" AND NOT "EStopAlarm";
   "Brake_Out" := ("BrakeHoa" = 1) OR (("BrakeHoa" = 2) AND "Brake_Ctrl");
   "AlarmHorn_Out" := ("AlarmHornHoa" = 1) OR (("AlarmHornHoa" = 2) AND "AlarmHorn_Ctrl");
   "StationInterlock_Out" := (("StationIntHoa" = 1) OR (("StationIntHoa" = 2) AND "StationIntl_Ctrl")) AND NOT "EStopAlarm";
   "Baffle_En" := ("BaffleHOA" = 1) OR (("BaffleHOA" = 2) AND "Baffle_Ctrl");
END_REGION

REGION Network 2
   // Analog Outputs
   RUNG wire#powerrail
      "SCP"(Input_Min := 0, Input_Signal := "OilPumpVFDpct", Input_Max := 100, Output_Min := 0, Output_Max := 27648, SV => "OilPumpVFDsp_Out")
   END_RUNG
   RUNG wire#powerrail
      "SCP"(Input_Min := 0, Input_Signal := "BafflePct", Input_Max := 100, Output_Min := 0, Output_Max := 27648, SV => "Baffle_Out")
   END_RUNG
   // the same network as SCL:
   "SCP"(Input_Min := 0,
         Input_Signal := "OilPumpVFDpct",
         Input_Max := 100,
         Output_Min := 0,
         Output_Max := 27648,
         SV => "OilPumpVFDsp_Out");
   "SCP"(Input_Min := 0,
         Input_Signal := "BafflePct",
         Input_Max := 100,
         Output_Min := 0,
         Output_Max := 27648,
         SV => "Baffle_Out");
END_REGION

REGION Network 3
   // Analog Inputs
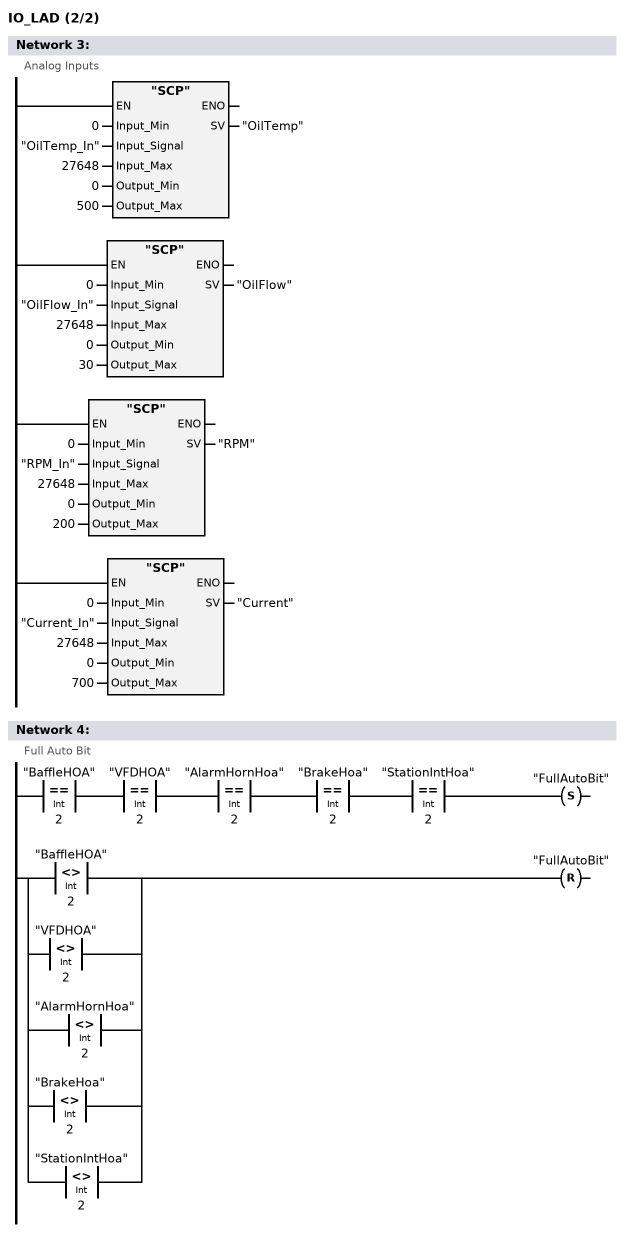
   RUNG wire#powerrail
      "SCP"(Input_Min := 0, Input_Signal := "OilTemp_In", Input_Max := 27648, Output_Min := 0, Output_Max := 500, SV => "OilTemp")
   END_RUNG
   RUNG wire#powerrail
      "SCP"(Input_Min := 0, Input_Signal := "OilFlow_In", Input_Max := 27648, Output_Min := 0, Output_Max := 30, SV => "OilFlow")
   END_RUNG
   RUNG wire#powerrail
      "SCP"(Input_Min := 0, Input_Signal := "RPM_In", Input_Max := 27648, Output_Min := 0, Output_Max := 200, SV => "RPM")
   END_RUNG
   RUNG wire#powerrail
      "SCP"(Input_Min := 0, Input_Signal := "Current_In", Input_Max := 27648, Output_Min := 0, Output_Max := 700, SV => "Current")
   END_RUNG
   // the same network as SCL:
   "SCP"(Input_Min := 0,
         Input_Signal := "OilTemp_In",
         Input_Max := 27648,
         Output_Min := 0,
         Output_Max := 500,
         SV => "OilTemp");
   "SCP"(Input_Min := 0,
         Input_Signal := "OilFlow_In",
         Input_Max := 27648,
         Output_Min := 0,
         Output_Max := 30,
         SV => "OilFlow");
   "SCP"(Input_Min := 0,
         Input_Signal := "RPM_In",
         Input_Max := 27648,
         Output_Min := 0,
         Output_Max := 200,
         SV => "RPM");
   "SCP"(Input_Min := 0,
         Input_Signal := "Current_In",
         Input_Max := 27648,
         Output_Min := 0,
         Output_Max := 700,
         SV => "Current");
END_REGION

REGION Network 4
   // Full Auto Bit
   RUNG wire#powerrail
      { S7_Templates := "SrcType := Int" } EQ_Contact(in1 := "BaffleHOA", in2 := 2)
      { S7_Templates := "SrcType := Int" } EQ_Contact(in1 := "VFDHOA", in2 := 2)
      { S7_Templates := "SrcType := Int" } EQ_Contact(in1 := "AlarmHornHoa", in2 := 2)
      { S7_Templates := "SrcType := Int" } EQ_Contact(in1 := "BrakeHoa", in2 := 2)
      { S7_Templates := "SrcType := Int" } EQ_Contact(in1 := "StationIntHoa", in2 := 2)
      S_Coil( "FullAutoBit" )
   END_RUNG
   RUNG wire#powerrail
      { S7_Templates := "SrcType := Int" } NE_Contact(in1 := "BaffleHOA", in2 := 2)
      wire#w1
      R_Coil( "FullAutoBit" )
   END_RUNG
   RUNG wire#powerrail
      { S7_Templates := "SrcType := Int" } NE_Contact(in1 := "VFDHOA", in2 := 2)
   END_RUNG wire#w1
   RUNG wire#powerrail
      { S7_Templates := "SrcType := Int" } NE_Contact(in1 := "AlarmHornHoa", in2 := 2)
   END_RUNG wire#w1
   RUNG wire#powerrail
      { S7_Templates := "SrcType := Int" } NE_Contact(in1 := "BrakeHoa", in2 := 2)
   END_RUNG wire#w1
   RUNG wire#powerrail
      { S7_Templates := "SrcType := Int" } NE_Contact(in1 := "StationIntHoa", in2 := 2)
   END_RUNG wire#w1
   // the same network as SCL:
   IF ("BaffleHOA" = 2) AND ("VFDHOA" = 2) AND ("AlarmHornHoa" = 2) AND ("BrakeHoa" = 2) AND ("StationIntHoa" = 2) THEN
       "FullAutoBit" := TRUE;
   END_IF;
   IF ("BaffleHOA" <> 2) OR ("VFDHOA" <> 2) OR ("AlarmHornHoa" <> 2) OR ("BrakeHoa" <> 2) OR ("StationIntHoa" <> 2) THEN
       "FullAutoBit" := FALSE;
   END_IF;
END_REGION
END_FUNCTION_BLOCK

FUNCTION_BLOCK "IO_FBD"   // FB3, FBD
{ S7_Optimized_Access := 'TRUE' }
VERSION : 0.1
   VAR_TEMP
      tv : Real;
   END_VAR
BEGIN

REGION Network 1
   // Digital Outputs
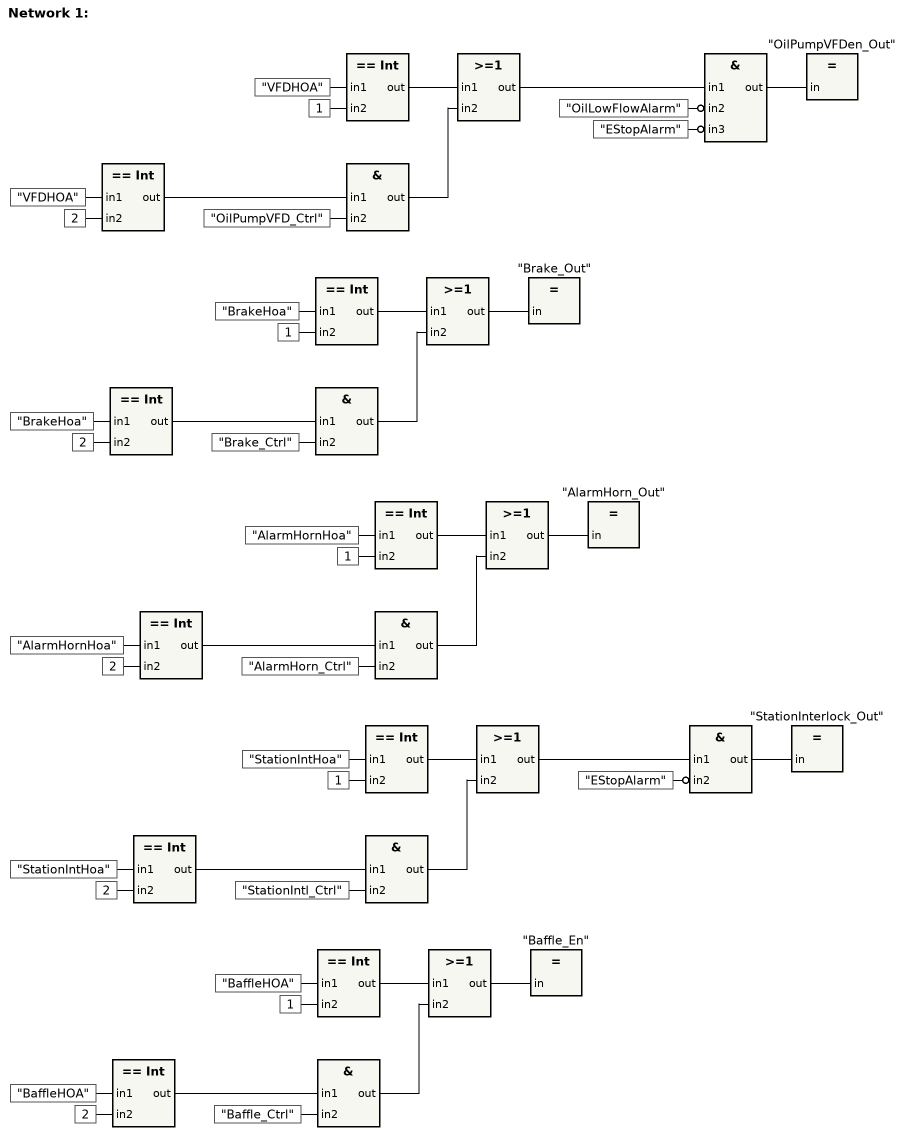
   "OilPumpVFDen_Out" := (("VFDHOA" = 1) OR (("VFDHOA" = 2) AND "OilPumpVFD_Ctrl")) AND NOT "OilLowFlowAlarm" AND NOT "EStopAlarm";
   "Brake_Out" := ("BrakeHoa" = 1) OR (("BrakeHoa" = 2) AND "Brake_Ctrl");
   "AlarmHorn_Out" := ("AlarmHornHoa" = 1) OR (("AlarmHornHoa" = 2) AND "AlarmHorn_Ctrl");
   "StationInterlock_Out" := (("StationIntHoa" = 1) OR (("StationIntHoa" = 2) AND "StationIntl_Ctrl")) AND NOT "EStopAlarm";
   "Baffle_En" := ("BaffleHOA" = 1) OR (("BaffleHOA" = 2) AND "Baffle_Ctrl");
END_REGION

REGION Network 2
   // Analog Outputs
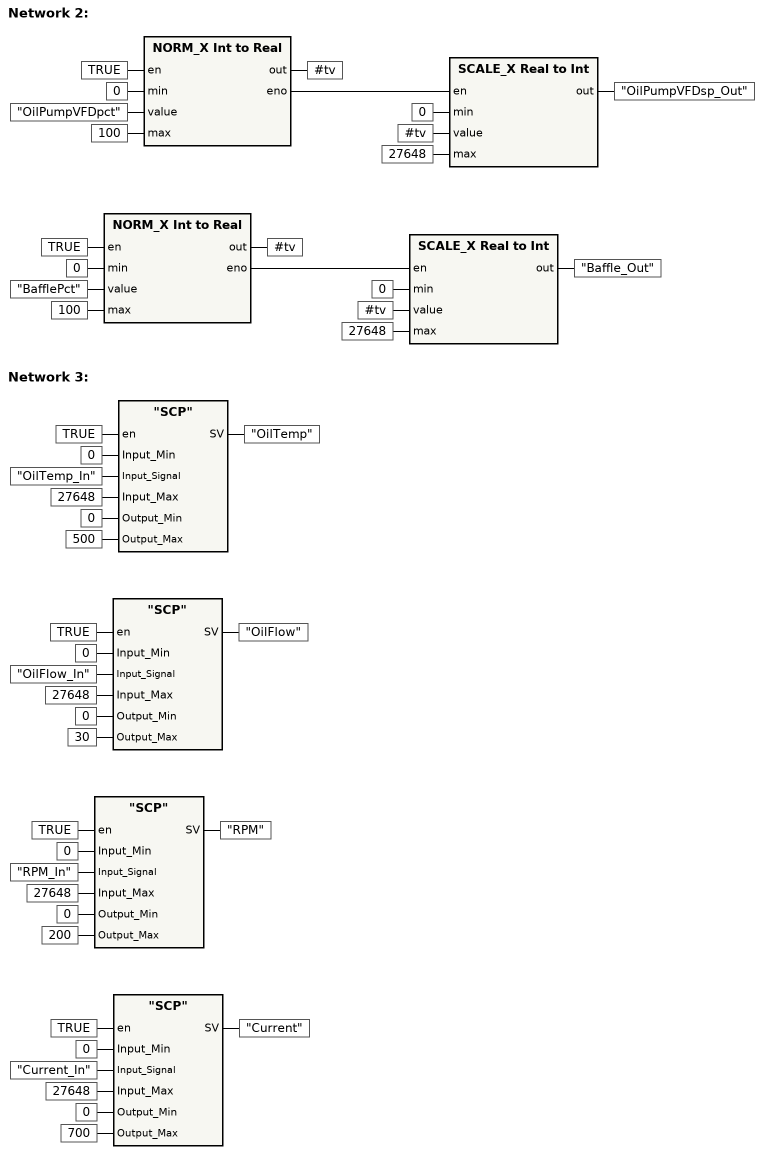
   IF TRUE THEN
       #tv := NORM_X(MIN := 0, VALUE := "OilPumpVFDpct", MAX := 100);
       "OilPumpVFDsp_Out" := SCALE_X(MIN := 0, VALUE := #tv, MAX := 27648);
       #tv := NORM_X(MIN := 0, VALUE := "BafflePct", MAX := 100);
       "Baffle_Out" := SCALE_X(MIN := 0, VALUE := #tv, MAX := 27648);
   END_IF;
END_REGION

REGION Network 3
   // Analog Inputs
   IF TRUE THEN
       "SCP"(Input_Min := 0,
             Input_Signal := "OilTemp_In",
             Input_Max := 27648,
             Output_Min := 0,
             Output_Max := 500,
             SV => "OilTemp");
       "SCP"(Input_Min := 0,
             Input_Signal := "OilFlow_In",
             Input_Max := 27648,
             Output_Min := 0,
             Output_Max := 30,
             SV => "OilFlow");
       "SCP"(Input_Min := 0,
             Input_Signal := "RPM_In",
             Input_Max := 27648,
             Output_Min := 0,
             Output_Max := 200,
             SV => "RPM");
       "SCP"(Input_Min := 0,
             Input_Signal := "Current_In",
             Input_Max := 27648,
             Output_Min := 0,
             Output_Max := 700,
             SV => "Current");
   END_IF;
END_REGION

REGION Network 4
   // Full Auto Bit
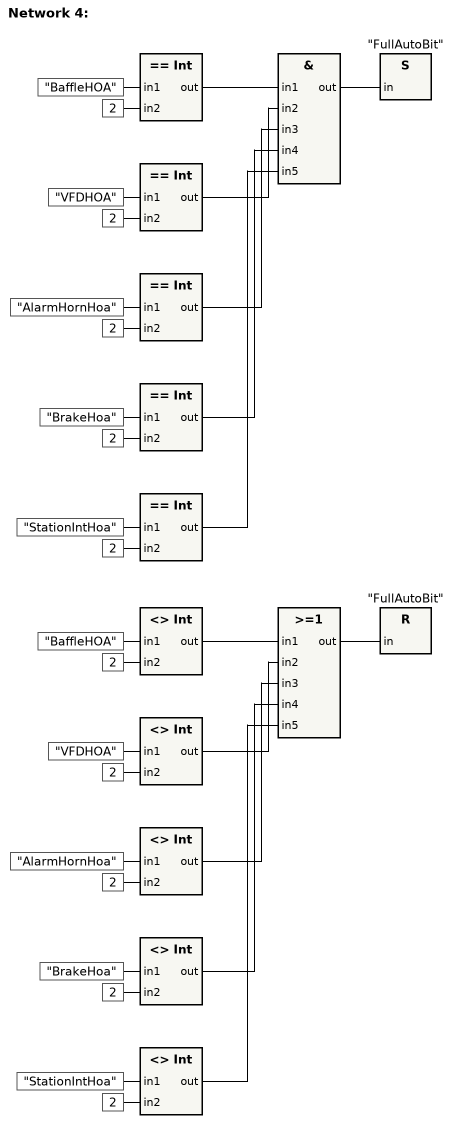
   IF ("BaffleHOA" = 2) AND ("VFDHOA" = 2) AND ("AlarmHornHoa" = 2) AND ("BrakeHoa" = 2) AND ("StationIntHoa" = 2) THEN
       "FullAutoBit" := TRUE;
   END_IF;
   IF ("BaffleHOA" <> 2) OR ("VFDHOA" <> 2) OR ("AlarmHornHoa" <> 2) OR ("BrakeHoa" <> 2) OR ("StationIntHoa" <> 2) THEN
       "FullAutoBit" := FALSE;
   END_IF;
END_REGION
END_FUNCTION_BLOCK

FUNCTION_BLOCK "IO_SCL"   // FB4, SCL
{ S7_Optimized_Access := 'TRUE' }
VERSION : 0.1
BEGIN
   //Digital Outputs
   IF "EStopAlarm" OR "OilLowFlowAlarm" OR "VFDHOA" = 0 OR ("VFDHOA" = 2 AND NOT "OilPumpVFD_Ctrl") THEN
       "OilPumpVFDen_Out" := 0;
   END_IF;

   IF ("VFDHOA" = 1 OR ("VFDHOA" = 2 AND "OilPumpVFD_Ctrl")) AND NOT "OilLowFlowAlarm" AND NOT "EStopAlarm" THEN
       "OilPumpVFDen_Out" := 1;
   END_IF;

   IF "BrakeHoa" = 0 OR ("BrakeHoa" = 2 AND NOT "Brake_Ctrl") THEN
       "Brake_Out" := 0;
   END_IF;

   IF "BrakeHoa" = 1 OR ("BrakeHoa" = 2 AND "Brake_Ctrl") THEN
       "Brake_Out" := 1;
   END_IF;

   IF "AlarmHornHoa" = 0 OR ("AlarmHornHoa" = 2 AND NOT "AlarmHorn_Ctrl") THEN
       "AlarmHorn_Out" := 0;
   END_IF;

   IF "AlarmHornHoa" = 1 OR ("AlarmHornHoa" = 2 AND "AlarmHorn_Ctrl") THEN
       "AlarmHorn_Out" := 1;
   END_IF;

   IF "StationIntHoa" = 0 OR ("StationIntHoa" = 2 AND NOT "StationIntl_Ctrl") THEN
       "StationInterlock_Out" := 0;
   END_IF;